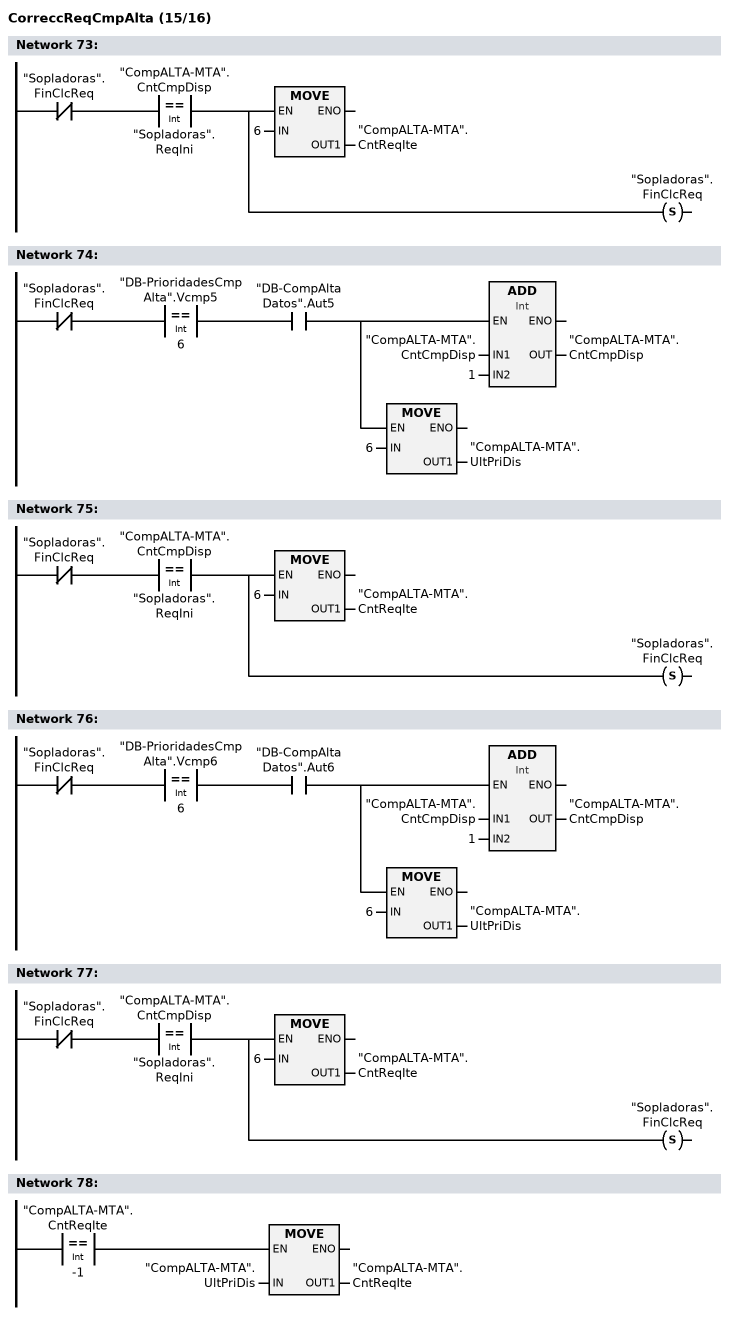
   RUNG wire#powerrail
      I_Contact( "Sopladoras".FinClcReq )
      { S7_Templates := "SrcType := Int" } EQ_Contact(in1 := "CompALTA-MTA".CntCmpDisp, in2 := "Sopladoras".ReqIni)
      wire#w1
      { S7_GenerateENO := "TRUE" } Move(in := 6, out1 => "CompALTA-MTA".CntReqIte)
   END_RUNG
   RUNG wire#w1
      S_Coil( "Sopladoras".FinClcReq )
   END_RUNG
   // the same network as SCL:
   IF NOT "Sopladoras".FinClcReq AND ("CompALTA-MTA".CntCmpDisp = "Sopladoras".ReqIni) THEN
       "CompALTA-MTA".CntReqIte := 6;
       "Sopladoras".FinClcReq := TRUE;
   END_IF;
END_REGION

REGION Network 74
   RUNG wire#powerrail
      I_Contact( "Sopladoras".FinClcReq )
      { S7_Templates := "SrcType := Int" } EQ_Contact(in1 := "DB-PrioridadesCmpAlta".Vcmp5, in2 := 6)
      Contact( "DB-CompAltaDatos".Aut5 )
      wire#w1
      { S7_Templates := "SrcType := Int"; S7_GenerateENO := "TRUE" } Add(in1 := "CompALTA-MTA".CntCmpDisp, in2 := 1, out => "CompALTA-MTA".CntCmpDisp)
   END_RUNG
   RUNG wire#w1
      { S7_GenerateENO := "TRUE" } Move(in := 6, out1 => "CompALTA-MTA".UltPriDis)
   END_RUNG
   // the same network as SCL:
   IF NOT "Sopladoras".FinClcReq AND ("DB-PrioridadesCmpAlta".Vcmp5 = 6) AND "DB-CompAltaDatos".Aut5 THEN
       "CompALTA-MTA".CntCmpDisp := "CompALTA-MTA".CntCmpDisp + 1;
       "CompALTA-MTA".UltPriDis := 6;
   END_IF;
END_REGION

REGION Network 75
   RUNG wire#powerrail
      I_Contact( "Sopladoras".FinClcReq )
      { S7_Templates := "SrcType := Int" } EQ_Contact(in1 := "CompALTA-MTA".CntCmpDisp, in2 := "Sopladoras".ReqIni)
      wire#w1
      { S7_GenerateENO := "TRUE" } Move(in := 6, out1 => "CompALTA-MTA".CntReqIte)
   END_RUNG
   RUNG wire#w1
      S_Coil( "Sopladoras".FinClcReq )
   END_RUNG
   // the same network as SCL:
   IF NOT "Sopladoras".FinClcReq AND ("CompALTA-MTA".CntCmpDisp = "Sopladoras".ReqIni) THEN
       "CompALTA-MTA".CntReqIte := 6;
       "Sopladoras".FinClcReq := TRUE;
   END_IF;
END_REGION

REGION Network 76
   RUNG wire#powerrail
      I_Contact( "Sopladoras".FinClcReq )
      { S7_Templates := "SrcType := Int" } EQ_Contact(in1 := "DB-PrioridadesCmpAlta".Vcmp6, in2 := 6)
      Contact( "DB-CompAltaDatos".Aut6 )
      wire#w1
      { S7_Templates := "SrcType := Int"; S7_GenerateENO := "TRUE" } Add(in1 := "CompALTA-MTA".CntCmpDisp, in2 := 1, out => "CompALTA-MTA".CntCmpDisp)
   END_RUNG
   RUNG wire#w1
      { S7_GenerateENO := "TRUE" } Move(in := 6, out1 => "CompALTA-MTA".UltPriDis)
   END_RUNG
   // the same network as SCL:
   IF NOT "Sopladoras".FinClcReq AND ("DB-PrioridadesCmpAlta".Vcmp6 = 6) AND "DB-CompAltaDatos".Aut6 THEN
       "CompALTA-MTA".CntCmpDisp := "CompALTA-MTA".CntCmpDisp + 1;
       "CompALTA-MTA".UltPriDis := 6;
   END_IF;
END_REGION

REGION Network 77
   RUNG wire#powerrail
      I_Contact( "Sopladoras".FinClcReq )
      { S7_Templates := "SrcType := Int" } EQ_Contact(in1 := "CompALTA-MTA".CntCmpDisp, in2 := "Sopladoras".ReqIni)
      wire#w1
      { S7_GenerateENO := "TRUE" } Move(in := 6, out1 => "CompALTA-MTA".CntReqIte)
   END_RUNG
   RUNG wire#w1
      S_Coil( "Sopladoras".FinClcReq )
   END_RUNG
   // the same network as SCL:
   IF NOT "Sopladoras".FinClcReq AND ("CompALTA-MTA".CntCmpDisp = "Sopladoras".ReqIni) THEN
       "CompALTA-MTA".CntReqIte := 6;
       "Sopladoras".FinClcReq := TRUE;
   END_IF;
END_REGION

REGION Network 78
   RUNG wire#powerrail
      { S7_Templates := "SrcType := Int" } EQ_Contact(in1 := "CompALTA-MTA".CntReqIte, in2 := -1)
      { S7_GenerateENO := "TRUE" } Move(in := "CompALTA-MTA".UltPriDis, out1 => "CompALTA-MTA".CntReqIte)
   END_RUNG
   // the same network as SCL:
   IF "CompALTA-MTA".CntReqIte = (-1) THEN "CompALTA-MTA".CntReqIte := "CompALTA-MTA".UltPriDis; END_IF;
END_REGION

REGION Network 79
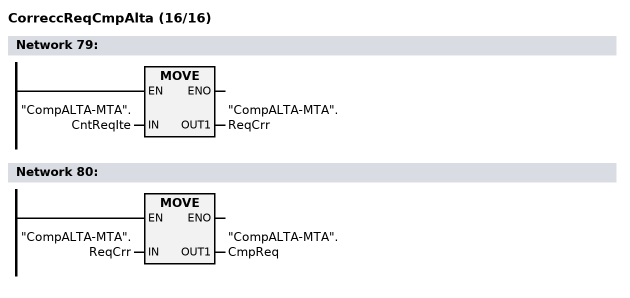
   RUNG wire#powerrail
      { S7_GenerateENO := "TRUE" } Move(in := "CompALTA-MTA".CntReqIte, out1 => "CompALTA-MTA".ReqCrr)
   END_RUNG
   // the same network as SCL:
   "CompALTA-MTA".ReqCrr := "CompALTA-MTA".CntReqIte;
END_REGION

REGION Network 80
   RUNG wire#powerrail
      { S7_GenerateENO := "TRUE" } Move(in := "CompALTA-MTA".ReqCrr, out1 => "CompALTA-MTA".CmpReq)
   END_RUNG
   // the same network as SCL:
   "CompALTA-MTA".CmpReq := "CompALTA-MTA".ReqCrr;
END_REGION
END_FUNCTION

FUNCTION "CalcEst6" : Void   // FC50, LAD
{ S7_Optimized_Access := 'FALSE' }
VERSION : 0.1
   VAR_TEMP   // added for the SCL form of the ladder/FBD networks
      _w1 : Bool;
   END_VAR
BEGIN

REGION Network 1: Prioritaria 1
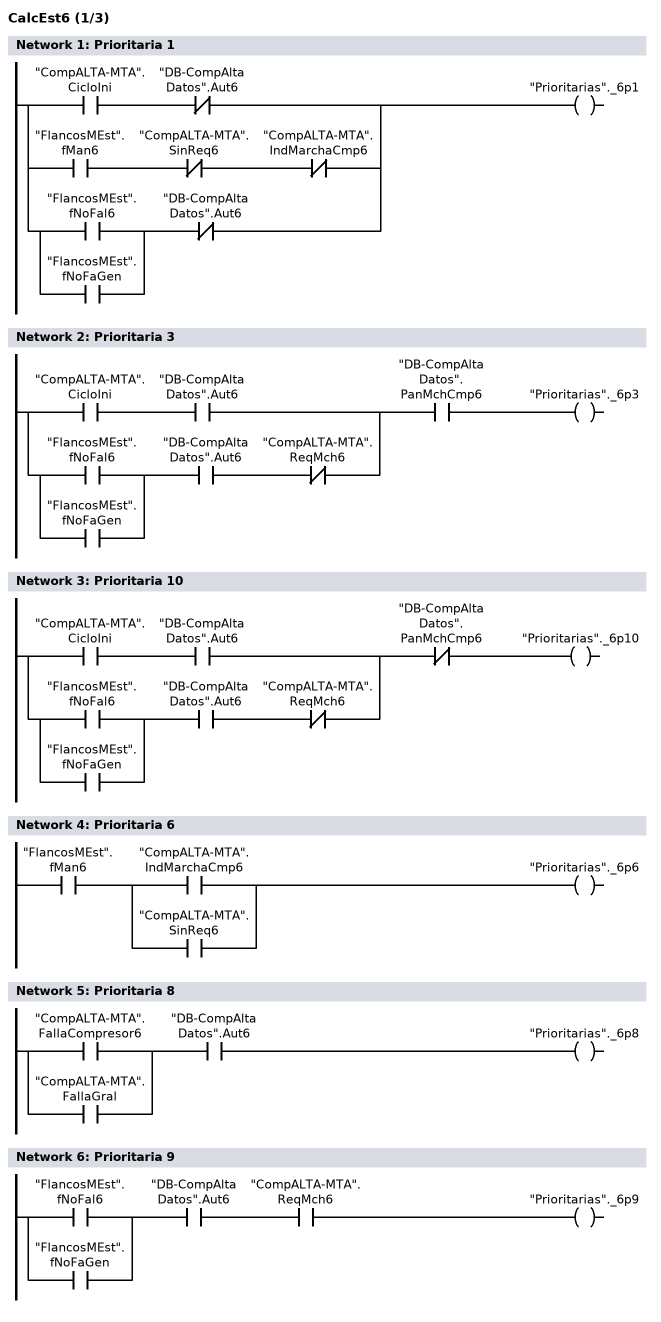
   RUNG wire#powerrail
      Contact( "CompALTA-MTA".CicloIni )
      I_Contact( "DB-CompAltaDatos".Aut6 )
      wire#w1
      Coil( "Prioritarias"._6p1 )
   END_RUNG
   RUNG wire#powerrail
      Contact( "FlancosMEst".fMan6 )
      I_Contact( "CompALTA-MTA".SinReq6 )
      I_Contact( "CompALTA-MTA".IndMarchaCmp6 )
   END_RUNG wire#w1
   RUNG wire#powerrail
      Contact( "FlancosMEst".fNoFal6 )
      wire#w2
      I_Contact( "DB-CompAltaDatos".Aut6 )
   END_RUNG wire#w1
   RUNG wire#powerrail
      Contact( "FlancosMEst".fNoFaGen )
   END_RUNG wire#w2
   // the same network as SCL:
   "Prioritarias"._6p1 := ("CompALTA-MTA".CicloIni AND NOT "DB-CompAltaDatos".Aut6) OR ("FlancosMEst".fMan6 AND NOT "CompALTA-MTA".SinReq6 AND NOT "CompALTA-MTA".IndMarchaCmp6) OR (("FlancosMEst".fNoFal6 OR "FlancosMEst".fNoFaGen) AND NOT "DB-CompAltaDatos".Aut6);
END_REGION

REGION Network 2: Prioritaria 3
   RUNG wire#powerrail
      Contact( "CompALTA-MTA".CicloIni )
      Contact( "DB-CompAltaDatos".Aut6 )
      wire#w1
      Contact( "DB-CompAltaDatos".PanMchCmp6 )
      Coil( "Prioritarias"._6p3 )
   END_RUNG
   RUNG wire#powerrail
      Contact( "FlancosMEst".fNoFal6 )
      wire#w2
      Contact( "DB-CompAltaDatos".Aut6 )
      I_Contact( "CompALTA-MTA".ReqMch6 )
   END_RUNG wire#w1
   RUNG wire#powerrail
      Contact( "FlancosMEst".fNoFaGen )
   END_RUNG wire#w2
   // the same network as SCL:
   "Prioritarias"._6p3 := (("CompALTA-MTA".CicloIni AND "DB-CompAltaDatos".Aut6) OR (("FlancosMEst".fNoFal6 OR "FlancosMEst".fNoFaGen) AND "DB-CompAltaDatos".Aut6 AND NOT "CompALTA-MTA".ReqMch6)) AND "DB-CompAltaDatos".PanMchCmp6;
END_REGION

REGION Network 3: Prioritaria 10
   RUNG wire#powerrail
      Contact( "CompALTA-MTA".CicloIni )
      Contact( "DB-CompAltaDatos".Aut6 )
      wire#w1
      I_Contact( "DB-CompAltaDatos".PanMchCmp6 )
      Coil( "Prioritarias"._6p10 )
   END_RUNG
   RUNG wire#powerrail
      Contact( "FlancosMEst".fNoFal6 )
      wire#w2
      Contact( "DB-CompAltaDatos".Aut6 )
      I_Contact( "CompALTA-MTA".ReqMch6 )
   END_RUNG wire#w1
   RUNG wire#powerrail
      Contact( "FlancosMEst".fNoFaGen )
   END_RUNG wire#w2
   // the same network as SCL:
   "Prioritarias"._6p10 := (("CompALTA-MTA".CicloIni AND "DB-CompAltaDatos".Aut6) OR (("FlancosMEst".fNoFal6 OR "FlancosMEst".fNoFaGen) AND "DB-CompAltaDatos".Aut6 AND NOT "CompALTA-MTA".ReqMch6)) AND NOT "DB-CompAltaDatos".PanMchCmp6;
END_REGION

REGION Network 4: Prioritaria 6
   RUNG wire#powerrail
      Contact( "FlancosMEst".fMan6 )
      wire#w1
      Contact( "CompALTA-MTA".IndMarchaCmp6 )
      wire#w2
      Coil( "Prioritarias"._6p6 )
   END_RUNG
   RUNG wire#w1
      Contact( "CompALTA-MTA".SinReq6 )
   END_RUNG wire#w2
   // the same network as SCL:
   "Prioritarias"._6p6 := "FlancosMEst".fMan6 AND ("CompALTA-MTA".IndMarchaCmp6 OR "CompALTA-MTA".SinReq6);
END_REGION

REGION Network 5: Prioritaria 8
   RUNG wire#powerrail
      Contact( "CompALTA-MTA".FallaCompresor6 )
      wire#w1
      Contact( "DB-CompAltaDatos".Aut6 )
      Coil( "Prioritarias"._6p8 )
   END_RUNG
   RUNG wire#powerrail
      Contact( "CompALTA-MTA".FallaGral )
   END_RUNG wire#w1
   // the same network as SCL:
   "Prioritarias"._6p8 := ("CompALTA-MTA".FallaCompresor6 OR "CompALTA-MTA".FallaGral) AND "DB-CompAltaDatos".Aut6;
END_REGION

REGION Network 6: Prioritaria 9
   RUNG wire#powerrail
      Contact( "FlancosMEst".fNoFal6 )
      wire#w1
      Contact( "DB-CompAltaDatos".Aut6 )
      Contact( "CompALTA-MTA".ReqMch6 )
      Coil( "Prioritarias"._6p9 )
   END_RUNG
   RUNG wire#powerrail
      Contact( "FlancosMEst".fNoFaGen )
   END_RUNG wire#w1
   // the same network as SCL:
   "Prioritarias"._6p9 := ("FlancosMEst".fNoFal6 OR "FlancosMEst".fNoFaGen) AND "DB-CompAltaDatos".Aut6 AND "CompALTA-MTA".ReqMch6;
END_REGION

REGION Network 7: Concatenadora 1
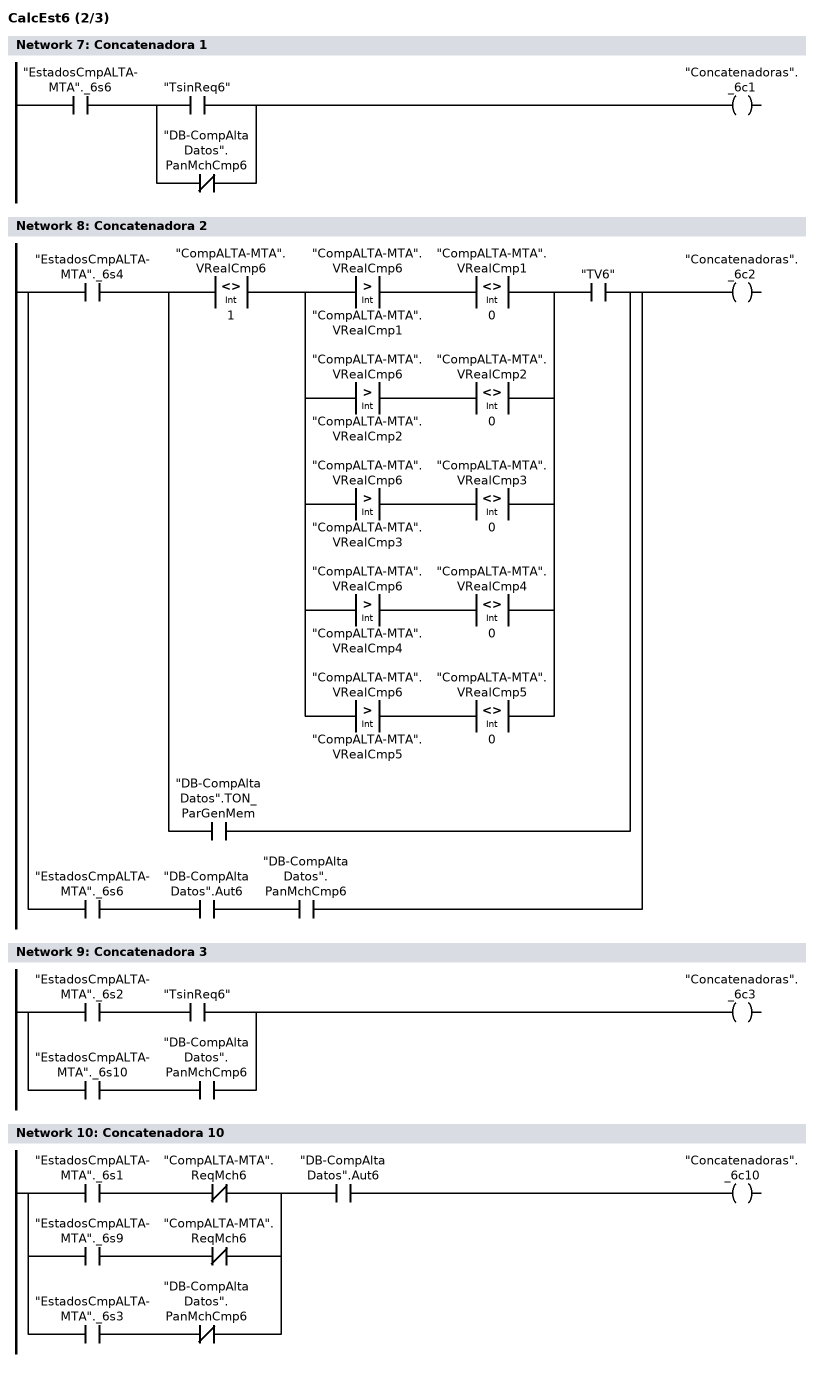
   RUNG wire#powerrail
      Contact( "EstadosCmpALTA-MTA"._6s6 )
      wire#w1
      Contact( "TsinReq6" )
      wire#w2
      Coil( "Concatenadoras"._6c1 )
   END_RUNG
   RUNG wire#w1
      I_Contact( "DB-CompAltaDatos".PanMchCmp6 )
   END_RUNG wire#w2
   // the same network as SCL:
   "Concatenadoras"._6c1 := "EstadosCmpALTA-MTA"._6s6 AND ("TsinReq6" OR NOT "DB-CompAltaDatos".PanMchCmp6);
END_REGION

REGION Network 8: Concatenadora 2
   RUNG wire#powerrail
      Contact( "EstadosCmpALTA-MTA"._6s4 )
      wire#w1
      { S7_Templates := "SrcType := Int" } NE_Contact(in1 := "CompALTA-MTA".VRealCmp6, in2 := 1)
      wire#w2
      { S7_Templates := "SrcType := Int" } GT_Contact(in1 := "CompALTA-MTA".VRealCmp6, in2 := "CompALTA-MTA".VRealCmp1)
      { S7_Templates := "SrcType := Int" } NE_Contact(in1 := "CompALTA-MTA".VRealCmp1, in2 := 0)
      wire#w3
      Contact( "TV6" )
      wire#w4
      Coil( "Concatenadoras"._6c2 )
   END_RUNG
   RUNG wire#w2
      { S7_Templates := "SrcType := Int" } GT_Contact(in1 := "CompALTA-MTA".VRealCmp6, in2 := "CompALTA-MTA".VRealCmp2)
      { S7_Templates := "SrcType := Int" } NE_Contact(in1 := "CompALTA-MTA".VRealCmp2, in2 := 0)
   END_RUNG wire#w3
   RUNG wire#w2
      { S7_Templates := "SrcType := Int" } GT_Contact(in1 := "CompALTA-MTA".VRealCmp6, in2 := "CompALTA-MTA".VRealCmp3)
      { S7_Templates := "SrcType := Int" } NE_Contact(in1 := "CompALTA-MTA".VRealCmp3, in2 := 0)
   END_RUNG wire#w3
   RUNG wire#w2
      { S7_Templates := "SrcType := Int" } GT_Contact(in1 := "CompALTA-MTA".VRealCmp6, in2 := "CompALTA-MTA".VRealCmp4)
      { S7_Templates := "SrcType := Int" } NE_Contact(in1 := "CompALTA-MTA".VRealCmp4, in2 := 0)
   END_RUNG wire#w3
   RUNG wire#w2
      { S7_Templates := "SrcType := Int" } GT_Contact(in1 := "CompALTA-MTA".VRealCmp6, in2 := "CompALTA-MTA".VRealCmp5)
      { S7_Templates := "SrcType := Int" } NE_Contact(in1 := "CompALTA-MTA".VRealCmp5, in2 := 0)
   END_RUNG wire#w3
   RUNG wire#w1
      Contact( "DB-CompAltaDatos".TON_ParGenMem )
   END_RUNG wire#w4
   RUNG wire#powerrail
      Contact( "EstadosCmpALTA-MTA"._6s6 )
      Contact( "DB-CompAltaDatos".Aut6 )
      Contact( "DB-CompAltaDatos".PanMchCmp6 )
   END_RUNG wire#w4
   // the same network as SCL:
   "Concatenadoras"._6c2 := ("EstadosCmpALTA-MTA"._6s4 AND ((("CompALTA-MTA".VRealCmp6 <> 1) AND ((("CompALTA-MTA".VRealCmp6 > "CompALTA-MTA".VRealCmp1) AND ("CompALTA-MTA".VRealCmp1 <> 0)) OR (("CompALTA-MTA".VRealCmp6 > "CompALTA-MTA".VRealCmp2) AND ("CompALTA-MTA".VRealCmp2 <> 0)) OR (("CompALTA-MTA".VRealCmp6 > "CompALTA-MTA".VRealCmp3) AND ("CompALTA-MTA".VRealCmp3 <> 0)) OR (("CompALTA-MTA".VRealCmp6 > "CompALTA-MTA".VRealCmp4) AND ("CompALTA-MTA".VRealCmp4 <> 0)) OR (("CompALTA-MTA".VRealCmp6 > "CompALTA-MTA".VRealCmp5) AND ("CompALTA-MTA".VRealCmp5 <> 0))) AND "TV6") OR "DB-CompAltaDatos".TON_ParGenMem)) OR ("EstadosCmpALTA-MTA"._6s6 AND "DB-CompAltaDatos".Aut6 AND "DB-CompAltaDatos".PanMchCmp6);
END_REGION

REGION Network 9: Concatenadora 3
   RUNG wire#powerrail
      Contact( "EstadosCmpALTA-MTA"._6s2 )
      Contact( "TsinReq6" )
      wire#w1
      Coil( "Concatenadoras"._6c3 )
   END_RUNG
   RUNG wire#powerrail
      Contact( "EstadosCmpALTA-MTA"._6s10 )
      Contact( "DB-CompAltaDatos".PanMchCmp6 )
   END_RUNG wire#w1
   // the same network as SCL:
   "Concatenadoras"._6c3 := ("EstadosCmpALTA-MTA"._6s2 AND "TsinReq6") OR ("EstadosCmpALTA-MTA"._6s10 AND "DB-CompAltaDatos".PanMchCmp6);
END_REGION

REGION Network 10: Concatenadora 10
   RUNG wire#powerrail
      Contact( "EstadosCmpALTA-MTA"._6s1 )
      I_Contact( "CompALTA-MTA".ReqMch6 )
      wire#w1
      Contact( "DB-CompAltaDatos".Aut6 )
      Coil( "Concatenadoras"._6c10 )
   END_RUNG
   RUNG wire#powerrail
      Contact( "EstadosCmpALTA-MTA"._6s9 )
      I_Contact( "CompALTA-MTA".ReqMch6 )
   END_RUNG wire#w1
   RUNG wire#powerrail
      Contact( "EstadosCmpALTA-MTA"._6s3 )
      I_Contact( "DB-CompAltaDatos".PanMchCmp6 )
   END_RUNG wire#w1
   // the same network as SCL:
   "Concatenadoras"._6c10 := (("EstadosCmpALTA-MTA"._6s1 AND NOT "CompALTA-MTA".ReqMch6) OR ("EstadosCmpALTA-MTA"._6s9 AND NOT "CompALTA-MTA".ReqMch6) OR ("EstadosCmpALTA-MTA"._6s3 AND NOT "DB-CompAltaDatos".PanMchCmp6)) AND "DB-CompAltaDatos".Aut6;
END_REGION

REGION Network 11: Concatenadora 4
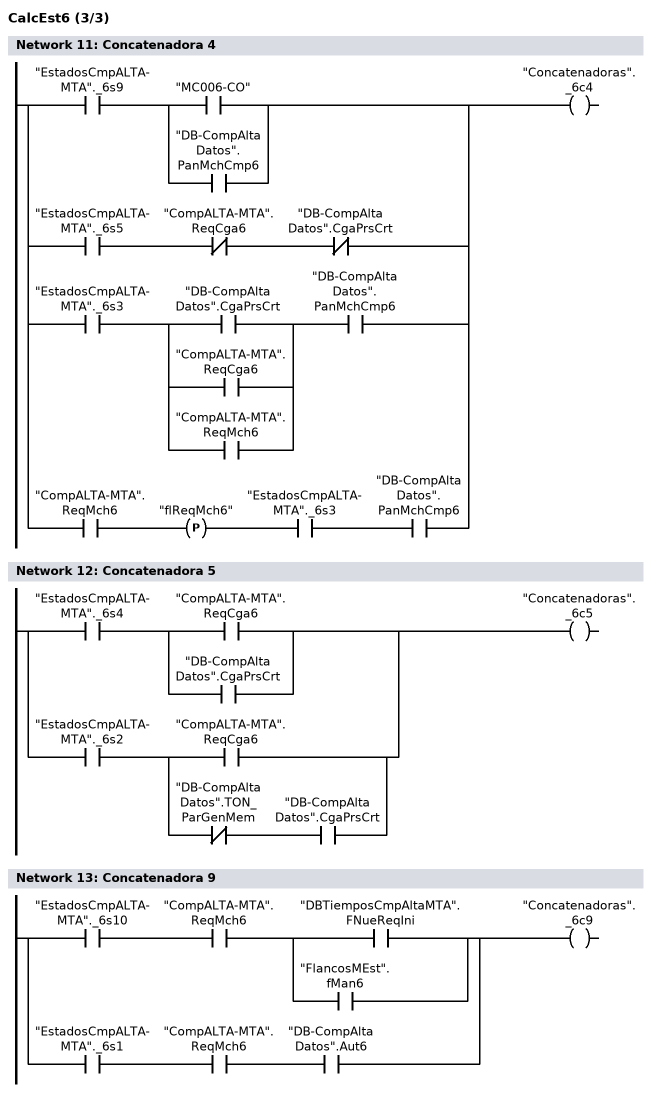
   RUNG wire#powerrail
      Contact( "EstadosCmpALTA-MTA"._6s9 )
      wire#w1
      Contact( "MC006-CO" )
      wire#w2
      Coil( "Concatenadoras"._6c4 )
   END_RUNG
   RUNG wire#w1
      Contact( "DB-CompAltaDatos".PanMchCmp6 )
   END_RUNG wire#w2
   RUNG wire#powerrail
      Contact( "EstadosCmpALTA-MTA"._6s5 )
      I_Contact( "CompALTA-MTA".ReqCga6 )
      I_Contact( "DB-CompAltaDatos".CgaPrsCrt )
   END_RUNG wire#w2
   RUNG wire#powerrail
      Contact( "EstadosCmpALTA-MTA"._6s3 )
      wire#w3
      Contact( "DB-CompAltaDatos".CgaPrsCrt )
      wire#w4
      Contact( "DB-CompAltaDatos".PanMchCmp6 )
   END_RUNG wire#w2
   RUNG wire#w3
      Contact( "CompALTA-MTA".ReqCga6 )
   END_RUNG wire#w4
   RUNG wire#w3
      Contact( "CompALTA-MTA".ReqMch6 )
   END_RUNG wire#w4
   RUNG wire#powerrail
      Contact( "CompALTA-MTA".ReqMch6 )
      P_Trig( "flReqMch6" )
      Contact( "EstadosCmpALTA-MTA"._6s3 )
      Contact( "DB-CompAltaDatos".PanMchCmp6 )
   END_RUNG wire#w2
   // the same network as SCL:
   #_w1 := "CompALTA-MTA".ReqMch6 AND NOT "flReqMch6";   // rising edge
   "flReqMch6" := "CompALTA-MTA".ReqMch6;
   "Concatenadoras"._6c4 := ("EstadosCmpALTA-MTA"._6s9 AND ("MC006-CO" OR "DB-CompAltaDatos".PanMchCmp6)) OR ("EstadosCmpALTA-MTA"._6s5 AND NOT "CompALTA-MTA".ReqCga6 AND NOT "DB-CompAltaDatos".CgaPrsCrt) OR ("EstadosCmpALTA-MTA"._6s3 AND ("DB-CompAltaDatos".CgaPrsCrt OR "CompALTA-MTA".ReqCga6 OR "CompALTA-MTA".ReqMch6) AND "DB-CompAltaDatos".PanMchCmp6) OR (#_w1 AND "EstadosCmpALTA-MTA"._6s3 AND "DB-CompAltaDatos".PanMchCmp6);
END_REGION

REGION Network 12: Concatenadora 5
   RUNG wire#powerrail
      Contact( "EstadosCmpALTA-MTA"._6s4 )
      wire#w1
      Contact( "CompALTA-MTA".ReqCga6 )
      wire#w2
      Coil( "Concatenadoras"._6c5 )
   END_RUNG
   RUNG wire#w1
      Contact( "DB-CompAltaDatos".CgaPrsCrt )
   END_RUNG wire#w2
   RUNG wire#powerrail
      Contact( "EstadosCmpALTA-MTA"._6s2 )
      wire#w3
      Contact( "CompALTA-MTA".ReqCga6 )
   END_RUNG wire#w2
   RUNG wire#w3
      I_Contact( "DB-CompAltaDatos".TON_ParGenMem )
      Contact( "DB-CompAltaDatos".CgaPrsCrt )
   END_RUNG wire#w2
   // the same network as SCL:
   "Concatenadoras"._6c5 := ("EstadosCmpALTA-MTA"._6s4 AND ("CompALTA-MTA".ReqCga6 OR "DB-CompAltaDatos".CgaPrsCrt)) OR ("EstadosCmpALTA-MTA"._6s2 AND ("CompALTA-MTA".ReqCga6 OR (NOT "DB-CompAltaDatos".TON_ParGenMem AND "DB-CompAltaDatos".CgaPrsCrt)));
END_REGION

REGION Network 13: Concatenadora 9
   RUNG wire#powerrail
      Contact( "EstadosCmpALTA-MTA"._6s10 )
      Contact( "CompALTA-MTA".ReqMch6 )
      wire#w1
      Contact( "DBTiemposCmpAltaMTA".FNueReqIni )
      wire#w2
      Coil( "Concatenadoras"._6c9 )
   END_RUNG
   RUNG wire#w1
      Contact( "FlancosMEst".fMan6 )
   END_RUNG wire#w2
   RUNG wire#powerrail
      Contact( "EstadosCmpALTA-MTA"._6s1 )
      Contact( "CompALTA-MTA".ReqMch6 )
      Contact( "DB-CompAltaDatos".Aut6 )
   END_RUNG wire#w2
   // the same network as SCL:
   "Concatenadoras"._6c9 := ("EstadosCmpALTA-MTA"._6s10 AND "CompALTA-MTA".ReqMch6 AND ("DBTiemposCmpAltaMTA".FNueReqIni OR "FlancosMEst".fMan6)) OR ("EstadosCmpALTA-MTA"._6s1 AND "CompALTA-MTA".ReqMch6 AND "DB-CompAltaDatos".Aut6);
END_REGION

REGION Network 14 (STL): Maquina de estados
         CALL  "FC_MAQ_EST_16"
         ( IN0  := %DB127.DBW10,
           IN1  := %DB128.DBW10,
           OUT2 := "ErrPMQ6",
           OUT3 := "ErrCMQ6",
           IO4  := %DB120.DBW10
         );
         NOP   0;
END_REGION

REGION Network 15 (STL): Bloque animación compresor
         CALL  "FC-ANIM-CMP"
         ( IN0  := %DB120.DBW10,
           OUT1 := "CompALTA-MTA".AnimCMP6
         );

         NOP   0;
END_REGION
END_FUNCTION

// folder: Compresores/Baja

FUNCTION "AutoCmpBaja" : Void   // FC24, LAD
{ S7_Optimized_Access := 'FALSE' }
VERSION : 0.1
   VAR_TEMP   // added for the SCL form of the ladder/FBD networks
      _w1 : Bool;
      _s5time1 : S5Time;
      _w2 : Bool;
   END_VAR
BEGIN

REGION Network 1 (STL)
         A(;
         L     "CmpBajaAuto".SPoffMC060;
         L     "CmpBajaAuto".SPonMC060;
         <=R;
         );
         JNB   M001;
         L     "CmpBajaAuto".SPonMC060;
         L     1;
         +R;
         T     "CmpBajaAuto".SPoffMC060;
   M001: NOP   0;
END_REGION

REGION Network 2 (STL)
         A(;
         L     "CmpBajaAuto".SPoffMC061;
         L     "CmpBajaAuto".SPonMC061;
         <=R;
         );
         JNB   M002;
         L     "CmpBajaAuto".SPonMC061;
         L     1;
         +R;
         T     "CmpBajaAuto".SPoffMC061;
   M002: NOP   0;
END_REGION

REGION Network 3 (STL)
         A(;
         L     "CmpBajaAuto".SPoffMC062;
         L     "CmpBajaAuto".SPonMC062;
         <=R;
         );
         JNB   M003;
         L     "CmpBajaAuto".SPonMC062;
         L     1;
         +R;
         T     "CmpBajaAuto".SPoffMC062;
   M003: NOP   0;
END_REGION

REGION Network 4 (STL)
         A(;
         L     "CmpBajaAuto".SPoffMC063;
         L     "CmpBajaAuto".SPonMC063;
         <=R;
         );
         JNB   M004;
         L     "CmpBajaAuto".SPonMC063;
         L     1;
         +R;
         T     "CmpBajaAuto".SPoffMC063;
   M004: NOP   0;
END_REGION

REGION Network 5 (STL)
         A(;
         L     "CmpBajaAuto".SPoffMC064;
         L     "CmpBajaAuto".SPonMC064;
         <=R;
         );
         JNB   M005;
         L     "CmpBajaAuto".SPonMC064;
         L     1;
         +R;
         T     "CmpBajaAuto".SPoffMC064;
   M005: NOP   0;
END_REGION

REGION Network 6
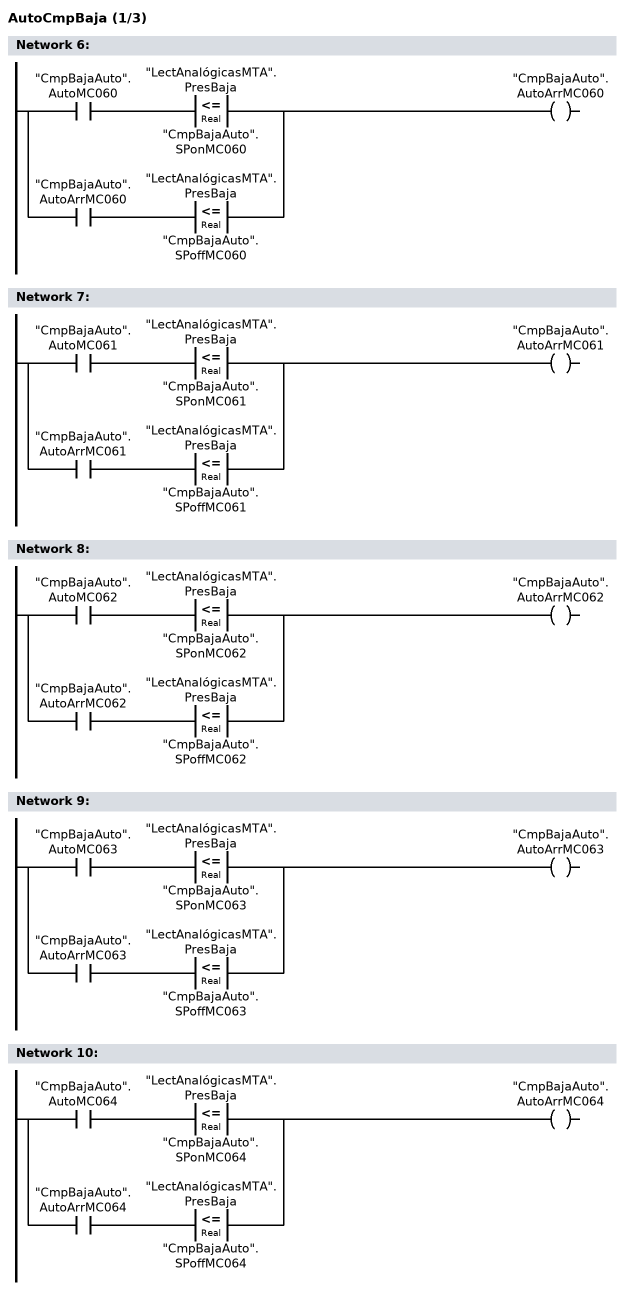
   "CmpBajaAuto".AutoArrMC060 := ("CmpBajaAuto".AutoMC060 AND ("LectAnalógicasMTA".PresBaja <= "CmpBajaAuto".SPonMC060)) OR ("CmpBajaAuto".AutoArrMC060 AND ("LectAnalógicasMTA".PresBaja <= "CmpBajaAuto".SPoffMC060));
END_REGION

REGION Network 7
   "CmpBajaAuto".AutoArrMC061 := ("CmpBajaAuto".AutoMC061 AND ("LectAnalógicasMTA".PresBaja <= "CmpBajaAuto".SPonMC061)) OR ("CmpBajaAuto".AutoArrMC061 AND ("LectAnalógicasMTA".PresBaja <= "CmpBajaAuto".SPoffMC061));
END_REGION

REGION Network 8
   "CmpBajaAuto".AutoArrMC062 := ("CmpBajaAuto".AutoMC062 AND ("LectAnalógicasMTA".PresBaja <= "CmpBajaAuto".SPonMC062)) OR ("CmpBajaAuto".AutoArrMC062 AND ("LectAnalógicasMTA".PresBaja <= "CmpBajaAuto".SPoffMC062));
END_REGION

REGION Network 9
   "CmpBajaAuto".AutoArrMC063 := ("CmpBajaAuto".AutoMC063 AND ("LectAnalógicasMTA".PresBaja <= "CmpBajaAuto".SPonMC063)) OR ("CmpBajaAuto".AutoArrMC063 AND ("LectAnalógicasMTA".PresBaja <= "CmpBajaAuto".SPoffMC063));
END_REGION

REGION Network 10
   "CmpBajaAuto".AutoArrMC064 := ("CmpBajaAuto".AutoMC064 AND ("LectAnalógicasMTA".PresBaja <= "CmpBajaAuto".SPonMC064)) OR ("CmpBajaAuto".AutoArrMC064 AND ("LectAnalógicasMTA".PresBaja <= "CmpBajaAuto".SPoffMC064));
END_REGION

REGION Network 11
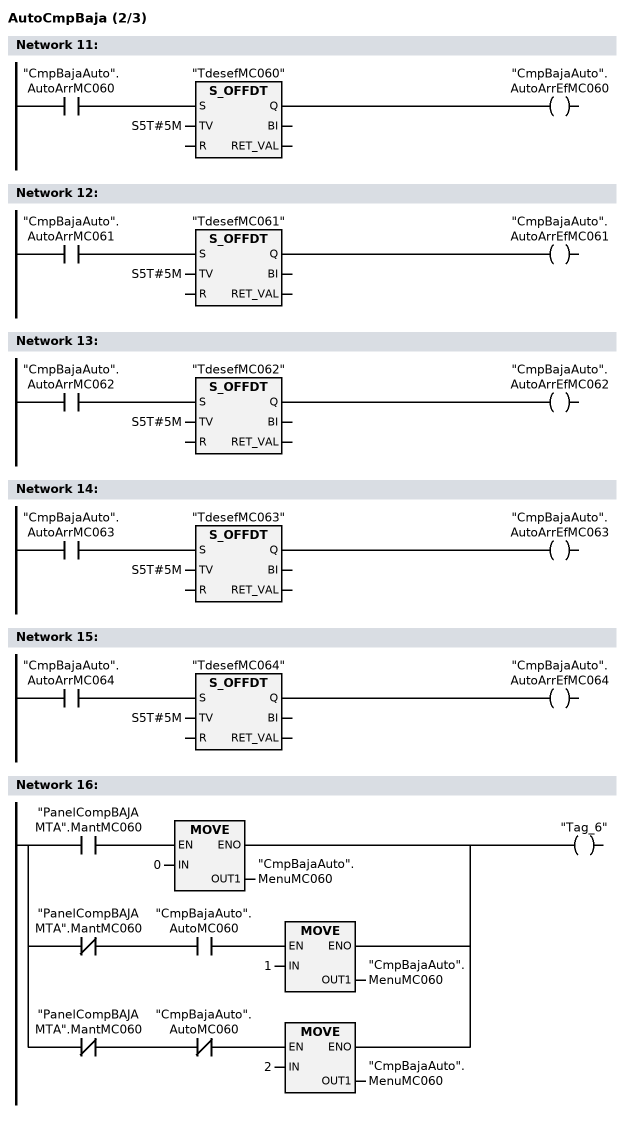
   RUNG wire#powerrail
      Contact( "CmpBajaAuto".AutoArrMC060 )
      S_OFFDT(T_NO := "TdesefMC060", TV := S5T#5M, R :=, BI =>, RET_VAL =>)
      Coil( "CmpBajaAuto".AutoArrEfMC060 )
   END_RUNG
   // the same network as SCL:
   #_s5time1 := S_OFFDT(T_NO := "TdesefMC060", TV := S5T#5M, S := "CmpBajaAuto".AutoArrMC060, Q => #_w1);
   "CmpBajaAuto".AutoArrEfMC060 := #_w1;
END_REGION

REGION Network 12
   RUNG wire#powerrail
      Contact( "CmpBajaAuto".AutoArrMC061 )
      S_OFFDT(T_NO := "TdesefMC061", TV := S5T#5M, R :=, BI =>, RET_VAL =>)
      Coil( "CmpBajaAuto".AutoArrEfMC061 )
   END_RUNG
   // the same network as SCL:
   #_s5time1 := S_OFFDT(T_NO := "TdesefMC061", TV := S5T#5M, S := "CmpBajaAuto".AutoArrMC061, Q => #_w1);
   "CmpBajaAuto".AutoArrEfMC061 := #_w1;
END_REGION

REGION Network 13
   RUNG wire#powerrail
      Contact( "CmpBajaAuto".AutoArrMC062 )
      S_OFFDT(T_NO := "TdesefMC062", TV := S5T#5M, R :=, BI =>, RET_VAL =>)
      Coil( "CmpBajaAuto".AutoArrEfMC062 )
   END_RUNG
   // the same network as SCL:
   #_s5time1 := S_OFFDT(T_NO := "TdesefMC062", TV := S5T#5M, S := "CmpBajaAuto".AutoArrMC062, Q => #_w1);
   "CmpBajaAuto".AutoArrEfMC062 := #_w1;
END_REGION

REGION Network 14
   RUNG wire#powerrail
      Contact( "CmpBajaAuto".AutoArrMC063 )
      S_OFFDT(T_NO := "TdesefMC063", TV := S5T#5M, R :=, BI =>, RET_VAL =>)
      Coil( "CmpBajaAuto".AutoArrEfMC063 )
   END_RUNG
   // the same network as SCL:
   #_s5time1 := S_OFFDT(T_NO := "TdesefMC063", TV := S5T#5M, S := "CmpBajaAuto".AutoArrMC063, Q => #_w1);
   "CmpBajaAuto".AutoArrEfMC063 := #_w1;
END_REGION

REGION Network 15
   RUNG wire#powerrail
      Contact( "CmpBajaAuto".AutoArrMC064 )
      S_OFFDT(T_NO := "TdesefMC064", TV := S5T#5M, R :=, BI =>, RET_VAL =>)
      Coil( "CmpBajaAuto".AutoArrEfMC064 )
   END_RUNG
   // the same network as SCL:
   #_s5time1 := S_OFFDT(T_NO := "TdesefMC064", TV := S5T#5M, S := "CmpBajaAuto".AutoArrMC064, Q => #_w1);
   "CmpBajaAuto".AutoArrEfMC064 := #_w1;
END_REGION

REGION Network 16
   RUNG wire#powerrail
      Contact( "PanelCompBAJA MTA".MantMC060 )
      { S7_GenerateENO := "TRUE" } Move(in := 0, out1 => "CmpBajaAuto".MenuMC060)
      wire#w1
      Coil( "Tag_6" )
   END_RUNG
   RUNG wire#powerrail
      I_Contact( "PanelCompBAJA MTA".MantMC060 )
      Contact( "CmpBajaAuto".AutoMC060 )
      { S7_GenerateENO := "TRUE" } Move(in := 1, out1 => "CmpBajaAuto".MenuMC060)
   END_RUNG wire#w1
   RUNG wire#powerrail
      I_Contact( "PanelCompBAJA MTA".MantMC060 )
      I_Contact( "CmpBajaAuto".AutoMC060 )
      { S7_GenerateENO := "TRUE" } Move(in := 2, out1 => "CmpBajaAuto".MenuMC060)
   END_RUNG wire#w1
   // the same network as SCL:
   // ENO of a box is taken as its EN; it also drops when the box reports an error
   IF "PanelCompBAJA MTA".MantMC060 THEN "CmpBajaAuto".MenuMC060 := 0; END_IF;
   #_w1 := NOT "PanelCompBAJA MTA".MantMC060 AND "CmpBajaAuto".AutoMC060;
   IF #_w1 THEN "CmpBajaAuto".MenuMC060 := 1; END_IF;
   #_w2 := NOT "PanelCompBAJA MTA".MantMC060 AND NOT "CmpBajaAuto".AutoMC060;
   IF #_w2 THEN "CmpBajaAuto".MenuMC060 := 2; END_IF;
   "Tag_6" := "PanelCompBAJA MTA".MantMC060 OR #_w1 OR #_w2;
END_REGION

REGION Network 17
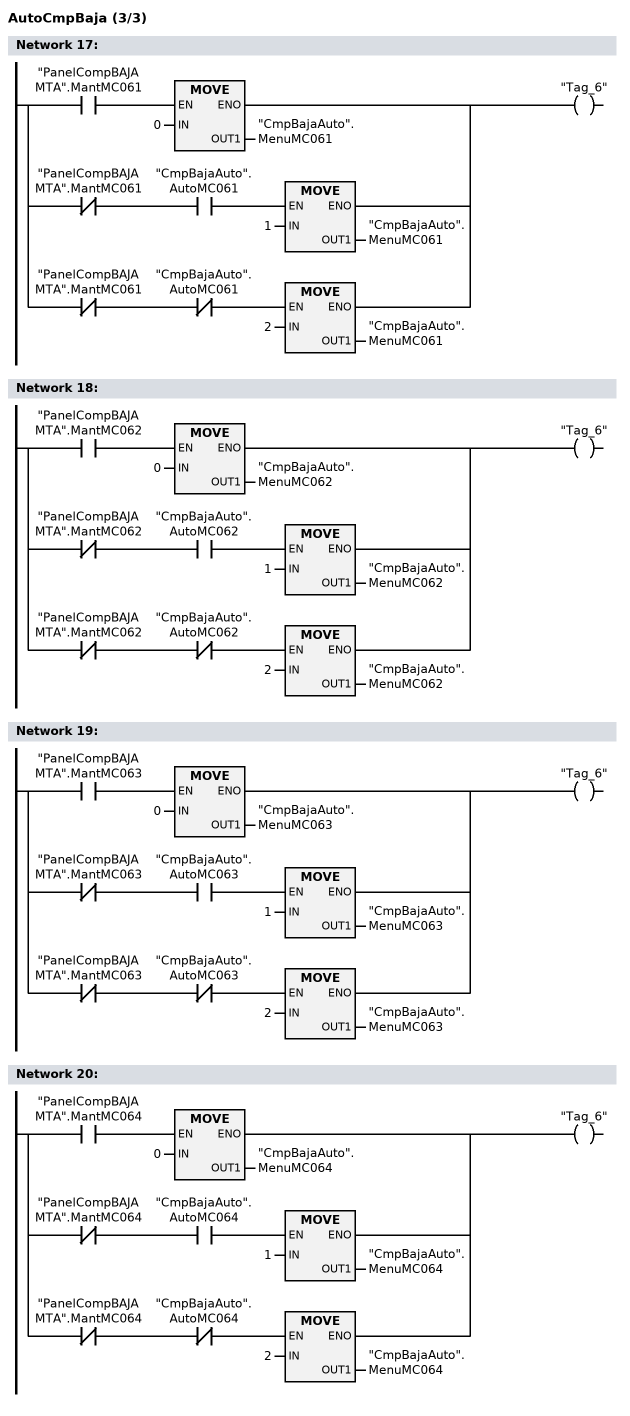
   RUNG wire#powerrail
      Contact( "PanelCompBAJA MTA".MantMC061 )
      { S7_GenerateENO := "TRUE" } Move(in := 0, out1 => "CmpBajaAuto".MenuMC061)
      wire#w1
      Coil( "Tag_6" )
   END_RUNG
   RUNG wire#powerrail
      I_Contact( "PanelCompBAJA MTA".MantMC061 )
      Contact( "CmpBajaAuto".AutoMC061 )
      { S7_GenerateENO := "TRUE" } Move(in := 1, out1 => "CmpBajaAuto".MenuMC061)
   END_RUNG wire#w1
   RUNG wire#powerrail
      I_Contact( "PanelCompBAJA MTA".MantMC061 )
      I_Contact( "CmpBajaAuto".AutoMC061 )
      { S7_GenerateENO := "TRUE" } Move(in := 2, out1 => "CmpBajaAuto".MenuMC061)
   END_RUNG wire#w1
   // the same network as SCL:
   // ENO of a box is taken as its EN; it also drops when the box reports an error
   IF "PanelCompBAJA MTA".MantMC061 THEN "CmpBajaAuto".MenuMC061 := 0; END_IF;
   #_w1 := NOT "PanelCompBAJA MTA".MantMC061 AND "CmpBajaAuto".AutoMC061;
   IF #_w1 THEN "CmpBajaAuto".MenuMC061 := 1; END_IF;
   #_w2 := NOT "PanelCompBAJA MTA".MantMC061 AND NOT "CmpBajaAuto".AutoMC061;
   IF #_w2 THEN "CmpBajaAuto".MenuMC061 := 2; END_IF;
   "Tag_6" := "PanelCompBAJA MTA".MantMC061 OR #_w1 OR #_w2;
END_REGION
